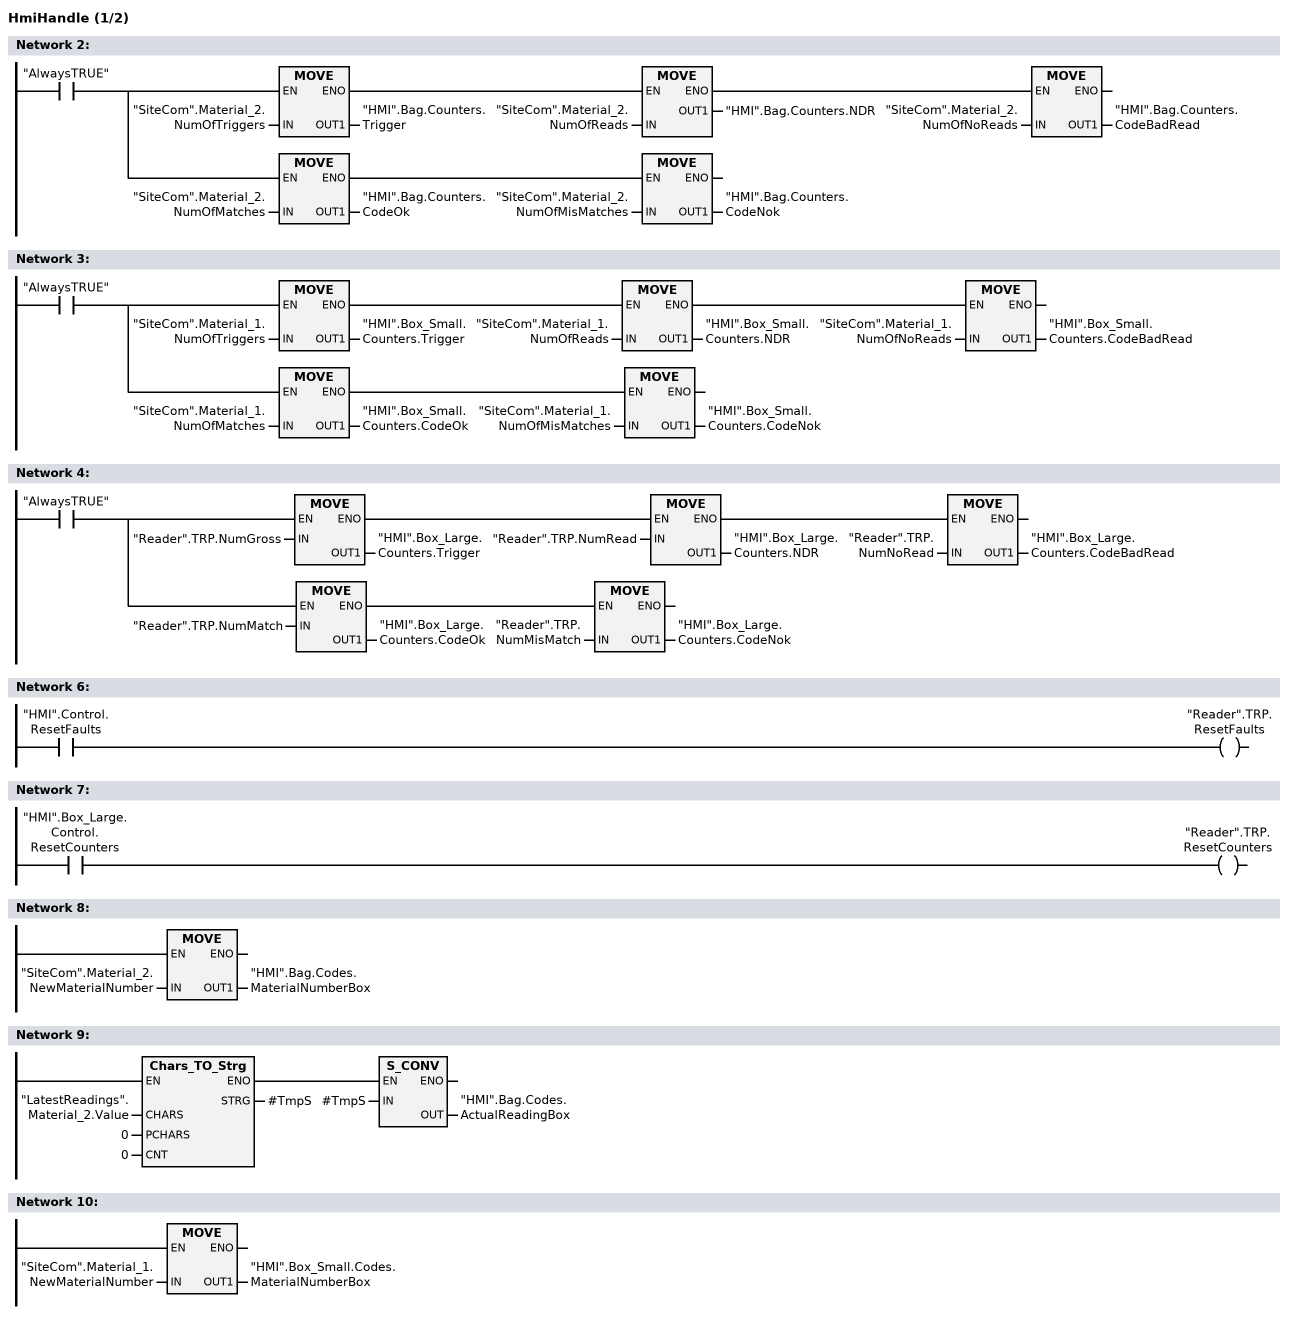
   RUNG wire#powerrail
      Contact( "AlwaysTRUE" )
      wire#w1
      Move(in := "SiteCom".Material_2.NumOfTriggers, out1 => "HMI".Bag.Counters.Trigger)
      Move(in := "SiteCom".Material_2.NumOfReads, out1 => "HMI".Bag.Counters.NDR)
      Move(in := "SiteCom".Material_2.NumOfNoReads, out1 => "HMI".Bag.Counters.CodeBadRead)
   END_RUNG
   RUNG wire#w1
      Move(in := "SiteCom".Material_2.NumOfMatches, out1 => "HMI".Bag.Counters.CodeOk)
      Move(in := "SiteCom".Material_2.NumOfMisMatches, out1 => "HMI".Bag.Counters.CodeNok)
   END_RUNG
   // the same network as SCL:
   IF "AlwaysTRUE" THEN
       "HMI".Bag.Counters.Trigger := "SiteCom".Material_2.NumOfTriggers;
       "HMI".Bag.Counters.NDR := "SiteCom".Material_2.NumOfReads;
       "HMI".Bag.Counters.CodeBadRead := "SiteCom".Material_2.NumOfNoReads;
       "HMI".Bag.Counters.CodeOk := "SiteCom".Material_2.NumOfMatches;
       "HMI".Bag.Counters.CodeNok := "SiteCom".Material_2.NumOfMisMatches;
   END_IF;
END_REGION

REGION Network 3
   RUNG wire#powerrail
      Contact( "AlwaysTRUE" )
      wire#w1
      Move(in := "SiteCom".Material_1.NumOfTriggers, out1 => "HMI".Box_Small.Counters.Trigger)
      Move(in := "SiteCom".Material_1.NumOfReads, out1 => "HMI".Box_Small.Counters.NDR)
      Move(in := "SiteCom".Material_1.NumOfNoReads, out1 => "HMI".Box_Small.Counters.CodeBadRead)
   END_RUNG
   RUNG wire#w1
      Move(in := "SiteCom".Material_1.NumOfMatches, out1 => "HMI".Box_Small.Counters.CodeOk)
      Move(in := "SiteCom".Material_1.NumOfMisMatches, out1 => "HMI".Box_Small.Counters.CodeNok)
   END_RUNG
   // the same network as SCL:
   IF "AlwaysTRUE" THEN
       "HMI".Box_Small.Counters.Trigger := "SiteCom".Material_1.NumOfTriggers;
       "HMI".Box_Small.Counters.NDR := "SiteCom".Material_1.NumOfReads;
       "HMI".Box_Small.Counters.CodeBadRead := "SiteCom".Material_1.NumOfNoReads;
       "HMI".Box_Small.Counters.CodeOk := "SiteCom".Material_1.NumOfMatches;
       "HMI".Box_Small.Counters.CodeNok := "SiteCom".Material_1.NumOfMisMatches;
   END_IF;
END_REGION

REGION Network 4
   RUNG wire#powerrail
      Contact( "AlwaysTRUE" )
      wire#w1
      Move(in := "Reader".TRP.NumGross, out1 => "HMI".Box_Large.Counters.Trigger)
      Move(in := "Reader".TRP.NumRead, out1 => "HMI".Box_Large.Counters.NDR)
      Move(in := "Reader".TRP.NumNoRead, out1 => "HMI".Box_Large.Counters.CodeBadRead)
   END_RUNG
   RUNG wire#w1
      Move(in := "Reader".TRP.NumMatch, out1 => "HMI".Box_Large.Counters.CodeOk)
      Move(in := "Reader".TRP.NumMisMatch, out1 => "HMI".Box_Large.Counters.CodeNok)
   END_RUNG
   // the same network as SCL:
   IF "AlwaysTRUE" THEN
       "HMI".Box_Large.Counters.Trigger := "Reader".TRP.NumGross;
       "HMI".Box_Large.Counters.NDR := "Reader".TRP.NumRead;
       "HMI".Box_Large.Counters.CodeBadRead := "Reader".TRP.NumNoRead;
       "HMI".Box_Large.Counters.CodeOk := "Reader".TRP.NumMatch;
       "HMI".Box_Large.Counters.CodeNok := "Reader".TRP.NumMisMatch;
   END_IF;
END_REGION

REGION Network 6
   RUNG wire#powerrail
      Contact( "HMI".Control.ResetFaults )
      Coil( "Reader".TRP.ResetFaults )
   END_RUNG
   // the same network as SCL:
   "Reader".TRP.ResetFaults := "HMI".Control.ResetFaults;
END_REGION

REGION Network 7
   RUNG wire#powerrail
      Contact( "HMI".Box_Large.Control.ResetCounters )
      Coil( "Reader".TRP.ResetCounters )
   END_RUNG
   // the same network as SCL:
   "Reader".TRP.ResetCounters := "HMI".Box_Large.Control.ResetCounters;
END_REGION

REGION Network 8
   RUNG wire#powerrail
      Move(in := "SiteCom".Material_2.NewMaterialNumber, out1 => "HMI".Bag.Codes.MaterialNumberBox)
   END_RUNG
   // the same network as SCL:
   "HMI".Bag.Codes.MaterialNumberBox := "SiteCom".Material_2.NewMaterialNumber;
END_REGION

REGION Network 9
   // no SCL statement known for Chars_TO_Strg: written as a call
   // ENO of a box is taken as its EN; it also drops when the box reports an error
   Chars_TO_Strg(Chars := "LatestReadings".Material_2.Value, pChars := 0, Cnt := 0, Strg => #TmpS);
   "HMI".Bag.Codes.ActualReadingBox := S_CONV(IN := #TmpS);
END_REGION

REGION Network 10
   RUNG wire#powerrail
      Move(in := "SiteCom".Material_1.NewMaterialNumber, out1 => "HMI".Box_Small.Codes.MaterialNumberBox)
   END_RUNG
   // the same network as SCL:
   "HMI".Box_Small.Codes.MaterialNumberBox := "SiteCom".Material_1.NewMaterialNumber;
END_REGION

REGION Network 11
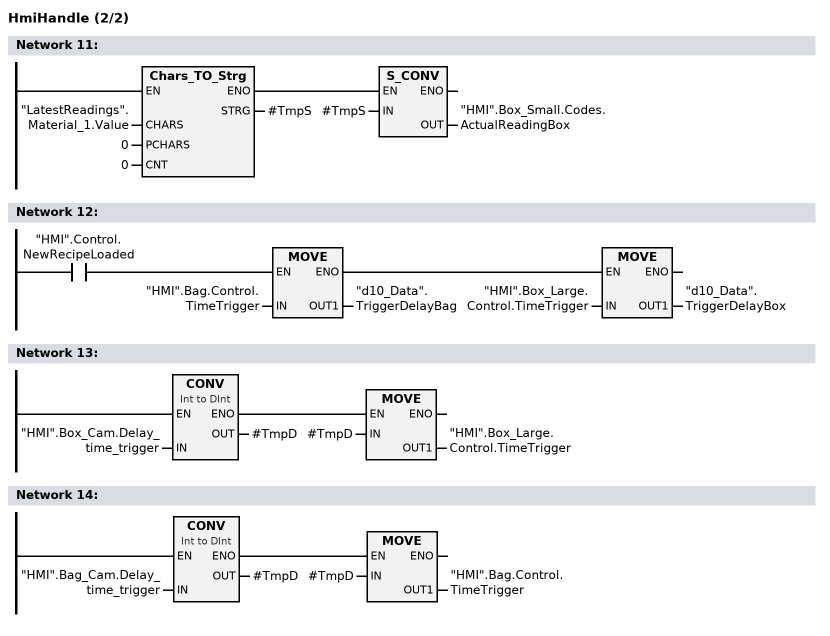
   // no SCL statement known for Chars_TO_Strg: written as a call
   // ENO of a box is taken as its EN; it also drops when the box reports an error
   Chars_TO_Strg(Chars := "LatestReadings".Material_1.Value, pChars := 0, Cnt := 0, Strg => #TmpS);
   "HMI".Box_Small.Codes.ActualReadingBox := S_CONV(IN := #TmpS);
END_REGION

REGION Network 12
   RUNG wire#powerrail
      Contact( "HMI".Control.NewRecipeLoaded )
      Move(in := "HMI".Bag.Control.TimeTrigger, out1 => "d10_Data".TriggerDelayBag)
      Move(in := "HMI".Box_Large.Control.TimeTrigger, out1 => "d10_Data".TriggerDelayBox)
   END_RUNG
   // the same network as SCL:
   IF "HMI".Control.NewRecipeLoaded THEN
       "d10_Data".TriggerDelayBag := "HMI".Bag.Control.TimeTrigger;
       "d10_Data".TriggerDelayBox := "HMI".Box_Large.Control.TimeTrigger;
   END_IF;
END_REGION

REGION Network 13
   RUNG wire#powerrail
      { S7_Templates := "[SrcType := Int, DestType := DInt]" } Convert(in := "HMI".Box_Cam.Delay_time_trigger, out => #TmpD)
      Move(in := #TmpD, out1 => "HMI".Box_Large.Control.TimeTrigger)
   END_RUNG
   // the same network as SCL:
   #TmpD := INT_TO_DINT("HMI".Box_Cam.Delay_time_trigger);
   "HMI".Box_Large.Control.TimeTrigger := #TmpD;
END_REGION

REGION Network 14
   RUNG wire#powerrail
      { S7_Templates := "[SrcType := Int, DestType := DInt]" } Convert(in := "HMI".Bag_Cam.Delay_time_trigger, out => #TmpD)
      Move(in := #TmpD, out1 => "HMI".Bag.Control.TimeTrigger)
   END_RUNG
   // the same network as SCL:
   #TmpD := INT_TO_DINT("HMI".Bag_Cam.Delay_time_trigger);
   "HMI".Bag.Control.TimeTrigger := #TmpD;
END_REGION
END_FUNCTION

FUNCTION "10_DataValidation" : Void   // FC10, LAD
{ S7_Optimized_Access := 'TRUE' }
VERSION : 0.1
BEGIN

REGION Network 1
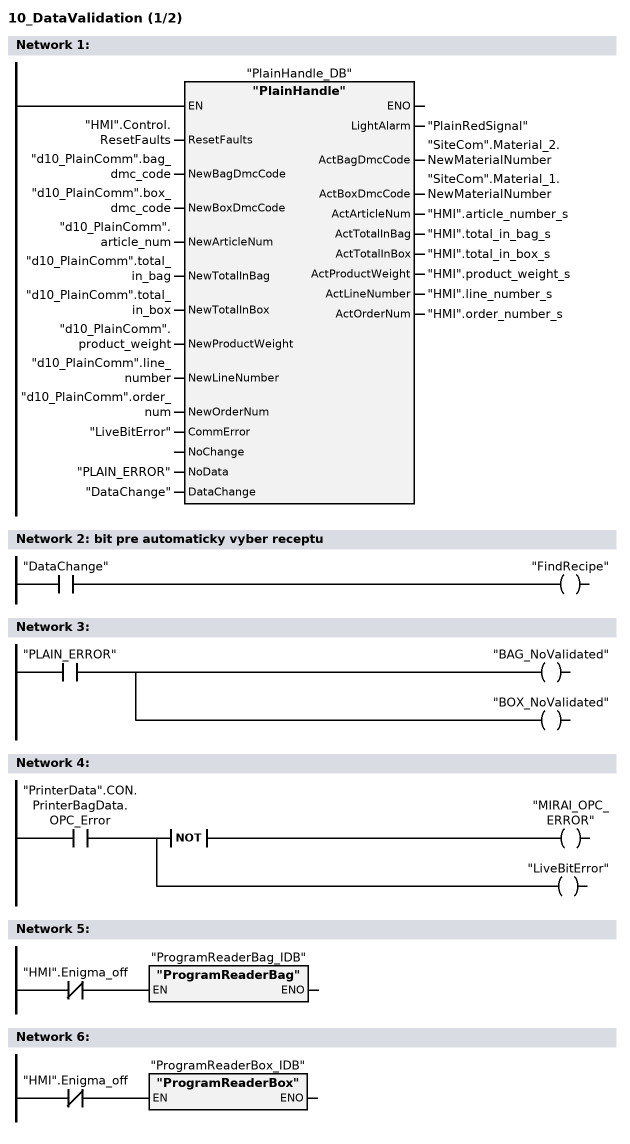
   RUNG wire#powerrail
      "PlainHandle_DB"(ResetFaults := "HMI".Control.ResetFaults, NewBagDmcCode := "d10_PlainComm".bag_dmc_code, NewBoxDmcCode := "d10_PlainComm".box_dmc_code, NewArticleNum := "d10_PlainComm".article_num, NewTotalInBag := "d10_PlainComm".total_in_bag, NewTotalInBox := "d10_PlainComm".total_in_box, NewProductWeight := "d10_PlainComm".product_weight, NewLineNumber := "d10_PlainComm".line_number, NewOrderNum := "d10_PlainComm".order_num, CommError := "LiveBitError", NoChange :=, NoData := "PLAIN_ERROR", DataChange := "DataChange", LightAlarm => "PlainRedSignal", ActBagDmcCode => "SiteCom".Material_2.NewMaterialNumber, ActBoxDmcCode => "SiteCom".Material_1.NewMaterialNumber, ActArticleNum => "HMI".article_number_s, ActTotalInBag => "HMI".total_in_bag_s, ActTotalInBox => "HMI".total_in_box_s, ActProductWeight => "HMI".product_weight_s, ActLineNumber => "HMI".line_number_s, ActOrderNum => "HMI".order_number_s)
   END_RUNG
   // the same network as SCL:
   "PlainHandle_DB"(ResetFaults := "HMI".Control.ResetFaults,   // "PlainHandle"
                    NewBagDmcCode := "d10_PlainComm".bag_dmc_code,
                    NewBoxDmcCode := "d10_PlainComm".box_dmc_code,
                    NewArticleNum := "d10_PlainComm".article_num,
                    NewTotalInBag := "d10_PlainComm".total_in_bag,
                    NewTotalInBox := "d10_PlainComm".total_in_box,
                    NewProductWeight := "d10_PlainComm".product_weight,
                    NewLineNumber := "d10_PlainComm".line_number,
                    NewOrderNum := "d10_PlainComm".order_num,
                    CommError := "LiveBitError",
                    NoData := "PLAIN_ERROR",
                    DataChange := "DataChange",
                    LightAlarm => "PlainRedSignal",
                    ActBagDmcCode => "SiteCom".Material_2.NewMaterialNumber,
                    ActBoxDmcCode => "SiteCom".Material_1.NewMaterialNumber,
                    ActArticleNum => "HMI".article_number_s,
                    ActTotalInBag => "HMI".total_in_bag_s,
                    ActTotalInBox => "HMI".total_in_box_s,
                    ActProductWeight => "HMI".product_weight_s,
                    ActLineNumber => "HMI".line_number_s,
                    ActOrderNum => "HMI".order_number_s);
END_REGION

REGION Network 2: bit pre automaticky vyber receptu
   RUNG wire#powerrail
      Contact( "DataChange" )
      Coil( "FindRecipe" )
   END_RUNG
   // the same network as SCL:
   "FindRecipe" := "DataChange";
END_REGION

REGION Network 3
   RUNG wire#powerrail
      Contact( "PLAIN_ERROR" )
      wire#w1
      Coil( "BAG_NoValidated" )
   END_RUNG
   RUNG wire#w1
      Coil( "BOX_NoValidated" )
   END_RUNG
   // the same network as SCL:
   "BAG_NoValidated" := "PLAIN_ERROR";
   "BOX_NoValidated" := "PLAIN_ERROR";
END_REGION

REGION Network 4
   RUNG wire#powerrail
      Contact( "PrinterData".CON.PrinterBagData.OPC_Error )
      wire#w1
      Not()
      Coil( "MIRAI_OPC_ERROR" )
   END_RUNG
   RUNG wire#w1
      Coil( "LiveBitError" )
   END_RUNG
   // the same network as SCL:
   "MIRAI_OPC_ERROR" := NOT "PrinterData".CON.PrinterBagData.OPC_Error;
   "LiveBitError" := "PrinterData".CON.PrinterBagData.OPC_Error;
END_REGION

REGION Network 5
   RUNG wire#powerrail
      I_Contact( "HMI".Enigma_off )
      "ProgramReaderBag_IDB"()
   END_RUNG
   // the same network as SCL:
   IF NOT "HMI".Enigma_off THEN
       "ProgramReaderBag_IDB"();   // "ProgramReaderBag"
   END_IF;
END_REGION

REGION Network 6
   RUNG wire#powerrail
      I_Contact( "HMI".Enigma_off )
      "ProgramReaderBox_IDB"()
   END_RUNG
   // the same network as SCL:
   IF NOT "HMI".Enigma_off THEN
       "ProgramReaderBox_IDB"();   // "ProgramReaderBox"
   END_IF;
END_REGION

REGION Network 7
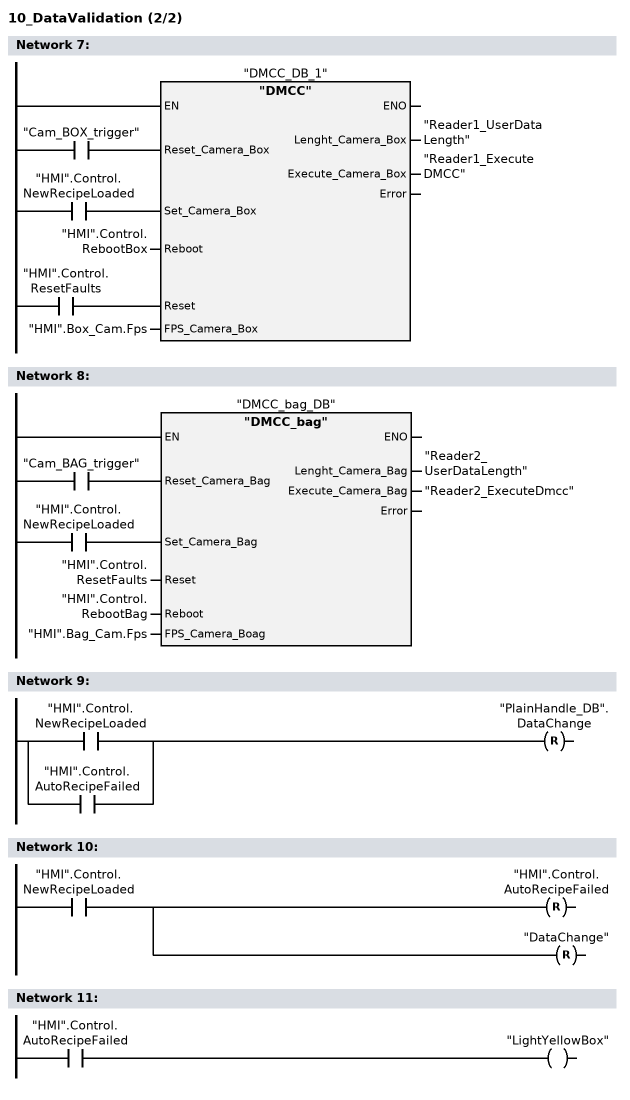
   RUNG wire#powerrail
      "DMCC_DB_1"(Reset_Camera_Box := wire#w1, Set_Camera_Box := wire#w2, Reset := wire#w3, Reboot := "HMI".Control.RebootBox, FPS_Camera_Box := "HMI".Box_Cam.Fps, Lenght_Camera_Box => "Reader1_UserData Length", Execute_Camera_Box => "Reader1_Execute DMCC", Error =>)
   END_RUNG
   RUNG wire#powerrail
      Contact( "Cam_BOX_trigger" )
   END_RUNG wire#w1
   RUNG wire#powerrail
      Contact( "HMI".Control.NewRecipeLoaded )
   END_RUNG wire#w2
   RUNG wire#powerrail
      Contact( "HMI".Control.ResetFaults )
   END_RUNG wire#w3
   // the same network as SCL:
   "DMCC_DB_1"(Reset_Camera_Box := "Cam_BOX_trigger",   // "DMCC"
               Set_Camera_Box := "HMI".Control.NewRecipeLoaded,
               Reboot := "HMI".Control.RebootBox,
               Reset := "HMI".Control.ResetFaults,
               FPS_Camera_Box := "HMI".Box_Cam.Fps,
               Lenght_Camera_Box => "Reader1_UserData Length",
               Execute_Camera_Box => "Reader1_Execute DMCC");
END_REGION

REGION Network 8
   RUNG wire#powerrail
      "DMCC_bag_DB"(Reset_Camera_Bag := wire#w1, Set_Camera_Bag := wire#w2, Reset := "HMI".Control.ResetFaults, Reboot := "HMI".Control.RebootBag, FPS_Camera_Boag := "HMI".Bag_Cam.Fps, Lenght_Camera_Bag => "Reader2_UserDataLength", Execute_Camera_Bag => "Reader2_ExecuteDmcc", Error =>)
   END_RUNG
   RUNG wire#powerrail
      Contact( "Cam_BAG_trigger" )
   END_RUNG wire#w1
   RUNG wire#powerrail
      Contact( "HMI".Control.NewRecipeLoaded )
   END_RUNG wire#w2
   // the same network as SCL:
   "DMCC_bag_DB"(Reset_Camera_Bag := "Cam_BAG_trigger",   // "DMCC_bag"
                 Set_Camera_Bag := "HMI".Control.NewRecipeLoaded,
                 Reset := "HMI".Control.ResetFaults,
                 Reboot := "HMI".Control.RebootBag,
                 FPS_Camera_Boag := "HMI".Bag_Cam.Fps,
                 Lenght_Camera_Bag => "Reader2_UserDataLength",
                 Execute_Camera_Bag => "Reader2_ExecuteDmcc");
END_REGION

REGION Network 9
   RUNG wire#powerrail
      Contact( "HMI".Control.NewRecipeLoaded )
      wire#w1
      R_Coil( "PlainHandle_DB".DataChange )
   END_RUNG
   RUNG wire#powerrail
      Contact( "HMI".Control.AutoRecipeFailed )
   END_RUNG wire#w1
   // the same network as SCL:
   IF "HMI".Control.NewRecipeLoaded OR "HMI".Control.AutoRecipeFailed THEN
       "PlainHandle_DB".DataChange := FALSE;
   END_IF;
END_REGION

REGION Network 10
   RUNG wire#powerrail
      Contact( "HMI".Control.NewRecipeLoaded )
      wire#w1
      R_Coil( "HMI".Control.AutoRecipeFailed )
   END_RUNG
   RUNG wire#w1
      R_Coil( "DataChange" )
   END_RUNG
   // the same network as SCL:
   IF "HMI".Control.NewRecipeLoaded THEN
       "HMI".Control.AutoRecipeFailed := FALSE;
       "DataChange" := FALSE;
   END_IF;
END_REGION

REGION Network 11
   RUNG wire#powerrail
      Contact( "HMI".Control.AutoRecipeFailed )
      Coil( "LightYellowBox" )
   END_RUNG
   // the same network as SCL:
   "LightYellowBox" := "HMI".Control.AutoRecipeFailed;
END_REGION
END_FUNCTION

FUNCTION "20_Mirai" : Void   // FC20, LAD
{ S7_Optimized_Access := 'TRUE' }
VERSION : 0.1
BEGIN

REGION Network 1
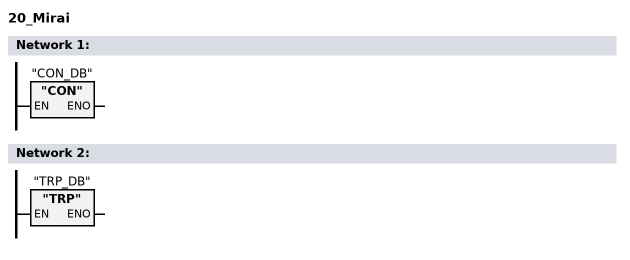
   RUNG wire#powerrail
      "CON_DB"()
   END_RUNG
   // the same network as SCL:
   "CON_DB"();   // "CON"
END_REGION

REGION Network 2
   RUNG wire#powerrail
      "TRP_DB"()
   END_RUNG
   // the same network as SCL:
   "TRP_DB"();   // "TRP"
END_REGION
END_FUNCTION

FUNCTION "FC_CleanQB_Bag" : Void   // FC100, LAD
{ S7_Optimized_Access := 'TRUE' }
VERSION : 0.1
BEGIN

REGION Network 1
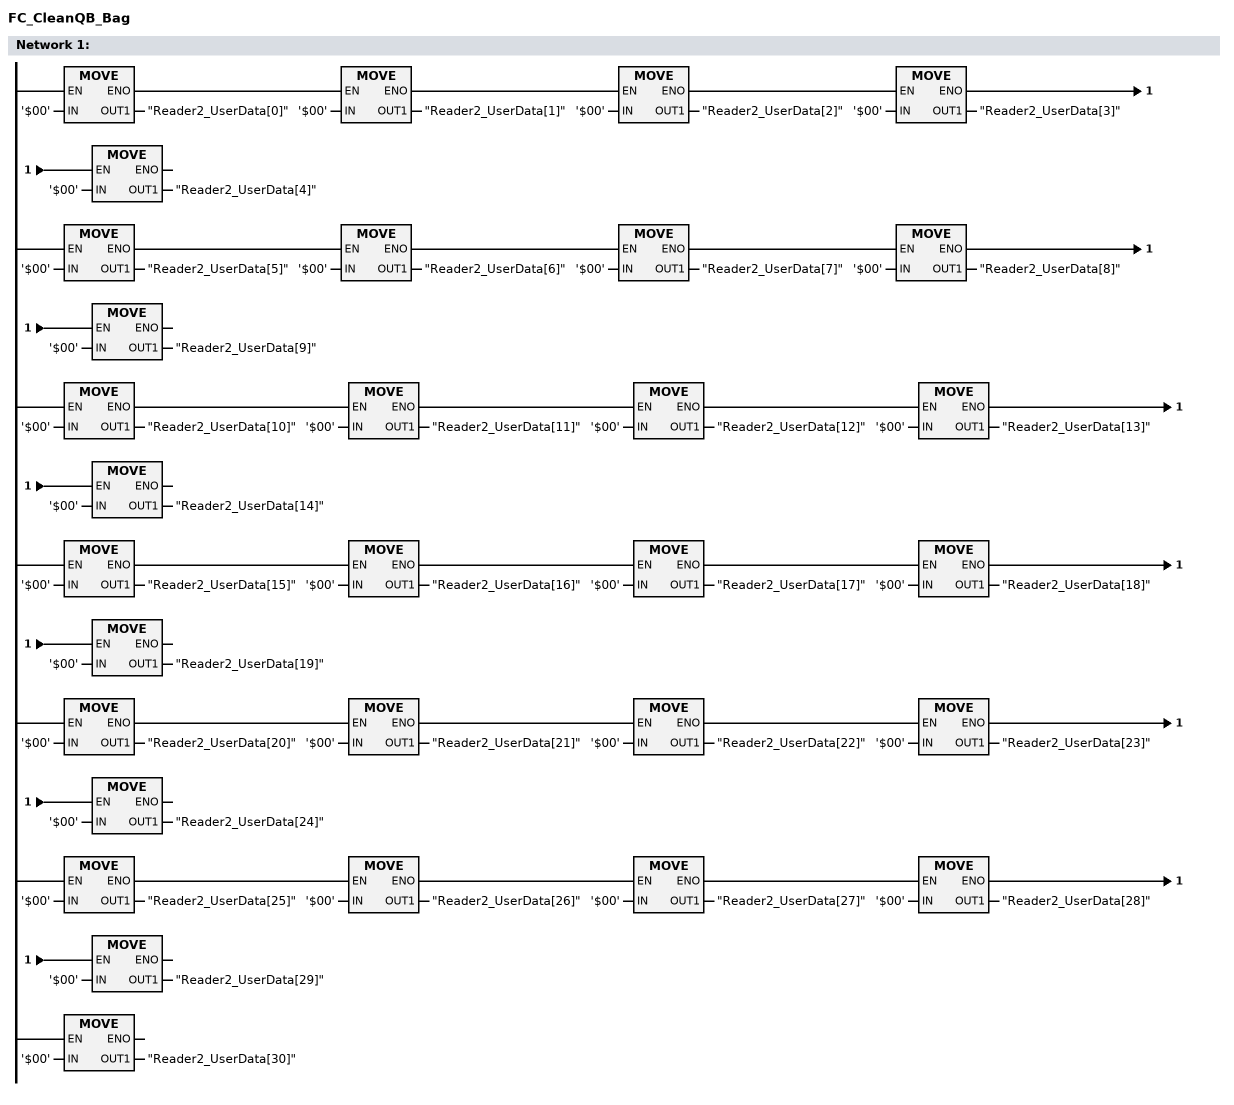
   RUNG wire#powerrail
      Move(in := '$00', out1 => "Reader2_UserData[0]")
      Move(in := '$00', out1 => "Reader2_UserData[1]")
      Move(in := '$00', out1 => "Reader2_UserData[2]")
      Move(in := '$00', out1 => "Reader2_UserData[3]")
      Move(in := '$00', out1 => "Reader2_UserData[4]")
   END_RUNG
   RUNG wire#powerrail
      Move(in := '$00', out1 => "Reader2_UserData[5]")
      Move(in := '$00', out1 => "Reader2_UserData[6]")
      Move(in := '$00', out1 => "Reader2_UserData[7]")
      Move(in := '$00', out1 => "Reader2_UserData[8]")
      Move(in := '$00', out1 => "Reader2_UserData[9]")
   END_RUNG
   RUNG wire#powerrail
      Move(in := '$00', out1 => "Reader2_UserData[10]")
      Move(in := '$00', out1 => "Reader2_UserData[11]")
      Move(in := '$00', out1 => "Reader2_UserData[12]")
      Move(in := '$00', out1 => "Reader2_UserData[13]")
      Move(in := '$00', out1 => "Reader2_UserData[14]")
   END_RUNG
   RUNG wire#powerrail
      Move(in := '$00', out1 => "Reader2_UserData[15]")
      Move(in := '$00', out1 => "Reader2_UserData[16]")
      Move(in := '$00', out1 => "Reader2_UserData[17]")
      Move(in := '$00', out1 => "Reader2_UserData[18]")
      Move(in := '$00', out1 => "Reader2_UserData[19]")
   END_RUNG
   RUNG wire#powerrail
      Move(in := '$00', out1 => "Reader2_UserData[20]")
      Move(in := '$00', out1 => "Reader2_UserData[21]")
      Move(in := '$00', out1 => "Reader2_UserData[22]")
      Move(in := '$00', out1 => "Reader2_UserData[23]")
      Move(in := '$00', out1 => "Reader2_UserData[24]")
   END_RUNG
   RUNG wire#powerrail
      Move(in := '$00', out1 => "Reader2_UserData[25]")
      Move(in := '$00', out1 => "Reader2_UserData[26]")
      Move(in := '$00', out1 => "Reader2_UserData[27]")
      Move(in := '$00', out1 => "Reader2_UserData[28]")
      Move(in := '$00', out1 => "Reader2_UserData[29]")
   END_RUNG
   RUNG wire#powerrail
      Move(in := '$00', out1 => "Reader2_UserData[30]")
   END_RUNG
   // the same network as SCL:
   "Reader2_UserData[0]" := '$00';
   "Reader2_UserData[1]" := '$00';
   "Reader2_UserData[2]" := '$00';
   "Reader2_UserData[3]" := '$00';
   "Reader2_UserData[4]" := '$00';
   "Reader2_UserData[5]" := '$00';
   "Reader2_UserData[6]" := '$00';
   "Reader2_UserData[7]" := '$00';
   "Reader2_UserData[8]" := '$00';
   "Reader2_UserData[9]" := '$00';
   "Reader2_UserData[10]" := '$00';
   "Reader2_UserData[11]" := '$00';
   "Reader2_UserData[12]" := '$00';
   "Reader2_UserData[13]" := '$00';
   "Reader2_UserData[14]" := '$00';
   "Reader2_UserData[15]" := '$00';
   "Reader2_UserData[16]" := '$00';
   "Reader2_UserData[17]" := '$00';
   "Reader2_UserData[18]" := '$00';
   "Reader2_UserData[19]" := '$00';
   "Reader2_UserData[20]" := '$00';
   "Reader2_UserData[21]" := '$00';
   "Reader2_UserData[22]" := '$00';
   "Reader2_UserData[23]" := '$00';
   "Reader2_UserData[24]" := '$00';
   "Reader2_UserData[25]" := '$00';
   "Reader2_UserData[26]" := '$00';
   "Reader2_UserData[27]" := '$00';
   "Reader2_UserData[28]" := '$00';
   "Reader2_UserData[29]" := '$00';
   "Reader2_UserData[30]" := '$00';
END_REGION
END_FUNCTION

FUNCTION "FC_CleanQB_Box" : Void   // FC101, LAD
{ S7_Optimized_Access := 'TRUE' }
VERSION : 0.1
BEGIN

REGION Network 1
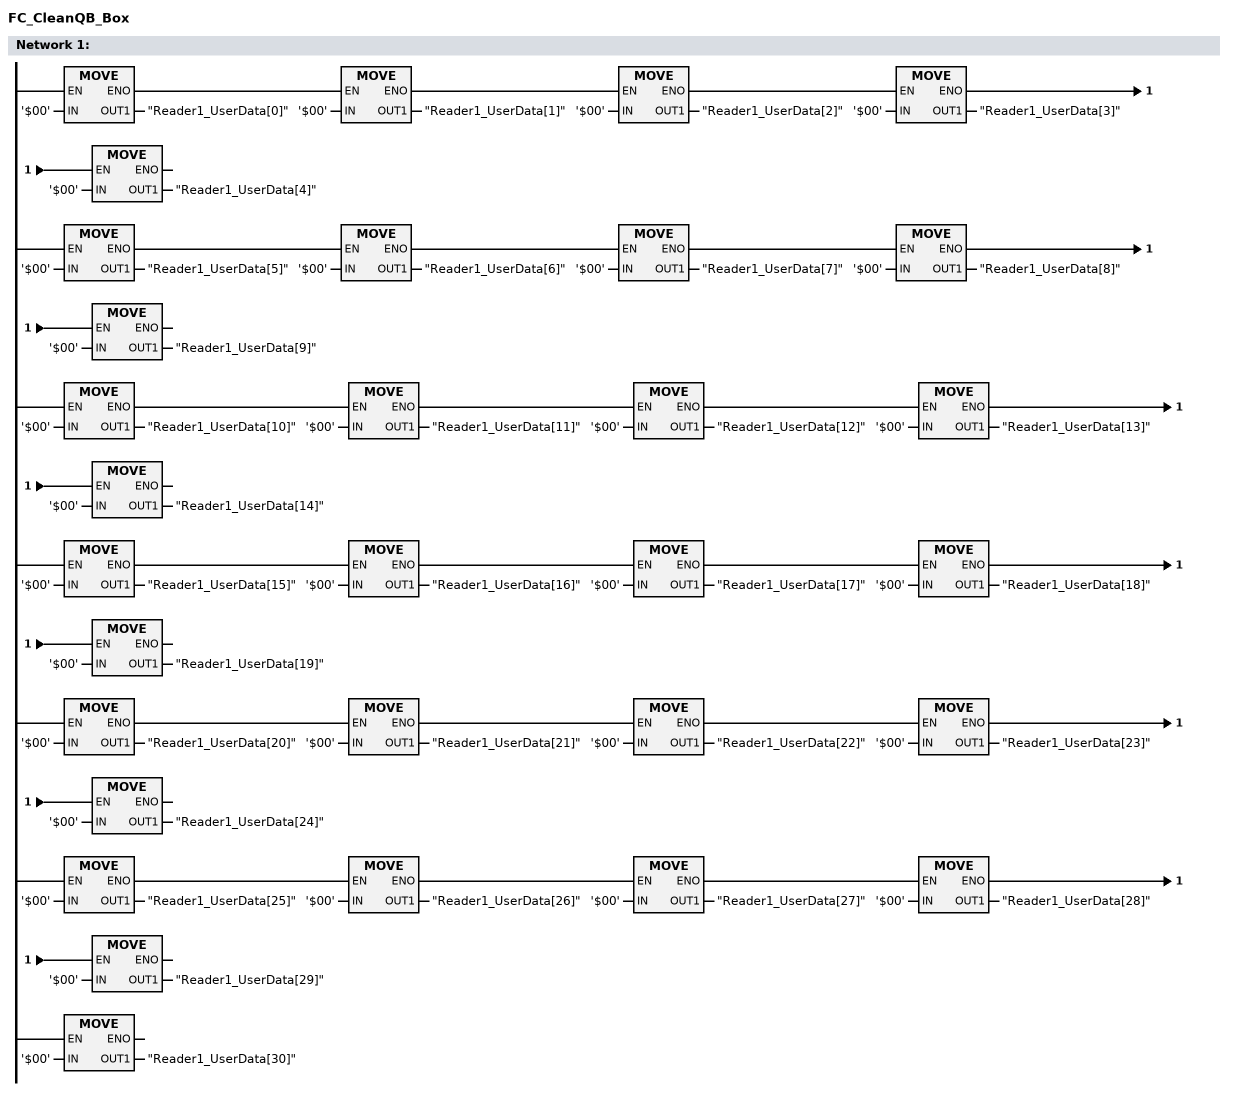
   RUNG wire#powerrail
      Move(in := '$00', out1 => "Reader1_UserData[0]")
      Move(in := '$00', out1 => "Reader1_UserData[1]")
      Move(in := '$00', out1 => "Reader1_UserData[2]")
      Move(in := '$00', out1 => "Reader1_UserData[3]")
      Move(in := '$00', out1 => "Reader1_UserData[4]")
   END_RUNG
   RUNG wire#powerrail
      Move(in := '$00', out1 => "Reader1_UserData[5]")
      Move(in := '$00', out1 => "Reader1_UserData[6]")
      Move(in := '$00', out1 => "Reader1_UserData[7]")
      Move(in := '$00', out1 => "Reader1_UserData[8]")
      Move(in := '$00', out1 => "Reader1_UserData[9]")
   END_RUNG
   RUNG wire#powerrail
      Move(in := '$00', out1 => "Reader1_UserData[10]")
      Move(in := '$00', out1 => "Reader1_UserData[11]")
      Move(in := '$00', out1 => "Reader1_UserData[12]")
      Move(in := '$00', out1 => "Reader1_UserData[13]")
      Move(in := '$00', out1 => "Reader1_UserData[14]")
   END_RUNG
   RUNG wire#powerrail
      Move(in := '$00', out1 => "Reader1_UserData[15]")
      Move(in := '$00', out1 => "Reader1_UserData[16]")
      Move(in := '$00', out1 => "Reader1_UserData[17]")
      Move(in := '$00', out1 => "Reader1_UserData[18]")
      Move(in := '$00', out1 => "Reader1_UserData[19]")
   END_RUNG
   RUNG wire#powerrail
      Move(in := '$00', out1 => "Reader1_UserData[20]")
      Move(in := '$00', out1 => "Reader1_UserData[21]")
      Move(in := '$00', out1 => "Reader1_UserData[22]")
      Move(in := '$00', out1 => "Reader1_UserData[23]")
      Move(in := '$00', out1 => "Reader1_UserData[24]")
   END_RUNG
   RUNG wire#powerrail
      Move(in := '$00', out1 => "Reader1_UserData[25]")
      Move(in := '$00', out1 => "Reader1_UserData[26]")
      Move(in := '$00', out1 => "Reader1_UserData[27]")
      Move(in := '$00', out1 => "Reader1_UserData[28]")
      Move(in := '$00', out1 => "Reader1_UserData[29]")
   END_RUNG
   RUNG wire#powerrail
      Move(in := '$00', out1 => "Reader1_UserData[30]")
   END_RUNG
   // the same network as SCL:
   "Reader1_UserData[0]" := '$00';
   "Reader1_UserData[1]" := '$00';
   "Reader1_UserData[2]" := '$00';
   "Reader1_UserData[3]" := '$00';
   "Reader1_UserData[4]" := '$00';
   "Reader1_UserData[5]" := '$00';
   "Reader1_UserData[6]" := '$00';
   "Reader1_UserData[7]" := '$00';
   "Reader1_UserData[8]" := '$00';
   "Reader1_UserData[9]" := '$00';
   "Reader1_UserData[10]" := '$00';
   "Reader1_UserData[11]" := '$00';
   "Reader1_UserData[12]" := '$00';
   "Reader1_UserData[13]" := '$00';
   "Reader1_UserData[14]" := '$00';
   "Reader1_UserData[15]" := '$00';
   "Reader1_UserData[16]" := '$00';
   "Reader1_UserData[17]" := '$00';
   "Reader1_UserData[18]" := '$00';
   "Reader1_UserData[19]" := '$00';
   "Reader1_UserData[20]" := '$00';
   "Reader1_UserData[21]" := '$00';
   "Reader1_UserData[22]" := '$00';
   "Reader1_UserData[23]" := '$00';
   "Reader1_UserData[24]" := '$00';
   "Reader1_UserData[25]" := '$00';
   "Reader1_UserData[26]" := '$00';
   "Reader1_UserData[27]" := '$00';
   "Reader1_UserData[28]" := '$00';
   "Reader1_UserData[29]" := '$00';
   "Reader1_UserData[30]" := '$00';
END_REGION
END_FUNCTION

FUNCTION "LGF_StringToTaddr" : TADDR_Param   // FC10041, SCL
{ S7_Optimized_Access := 'TRUE' }
VERSION : 0.1
   VAR_INPUT
      ipAddressString : String;
   END_VAR
   VAR_OUTPUT
      error : Bool;
      status : Word;
   END_VAR
   VAR_TEMP
      tempCharPosition : Int;
      tempAddressString : String;
      tempOctetString : String[4];
      tempUInt : UInt;
      tempPortNumberIsSpecified : Bool;
      tempIpAdressTaddr : TADDR_Param;
   END_VAR
   VAR CONSTANT
      NO_ERROR : Word := 16#0000;
      WRONG_VALUE_POS1 : Word := 16#8101;
      WRONG_VALUE_POS2 : Word := 16#8102;
      WRONG_VALUE_POS3 : Word := 16#8103;
      WRONG_VALUE_POS4 : Word := 16#8104;
      WRONG_VALUE_PORT : Word := 16#8105;
      MAX_USINT : USInt := 255;
      MAX_UINT : UInt := 65535;
      EMPTY_STRING : String := '';
      MAX_CHAR_FOR_IP_PART : Int := 4;
      MAX_CHAR_FOR_PORT_PART : Int := 5;
      INIT_VAL : USInt := 0;
      NO_POS : Int := 0;
   END_VAR
BEGIN
   //=============================================================================
   // SIEMENS AG
   // (c)Copyright 2017
   //-----------------------------------------------------------------------------
   // Library:       LGF (Library General Functions)
   // Tested with:   CPU1212C DC/DC/DC FW:V4.2
   // Engineering:   TIA Portal V14 Upd 1
   // Restrictions:  -
   // Requirements:  PLC (S7-1200 / S7-1500)
   // Functionality: This function converts a string IP Address
   //                into TADDR Param format.
   //-----------------------------------------------------------------------------
   // Change log table:
   // Version  Date       In charge Changes applied
   // 01.00.00 30.01.2017 Siemens Industry Online Support
   //                     First released version
   //-----------------------------------------------------------------------------
   //Status Codes:
   // 16#0000:  No errors
   // 16#8101:  Wrong value on position 1
   // 16#8102:  Wrong value on position 2
   // 16#8103:  Wrong value on position 3
   // 16#8104:  Wrong value on position 4
   // 16#8105:  Wrong value on port position
   //=============================================================================

   // Initialization
   #error := FALSE;
   #status := #NO_ERROR;
   #tempAddressString := #ipAddressString;
   #LGF_StringToTaddr.REM_IP_ADDR[1] := #INIT_VAL;
   #LGF_StringToTaddr.REM_IP_ADDR[2] := #INIT_VAL;
   #LGF_StringToTaddr.REM_IP_ADDR[3] := #INIT_VAL;
   #LGF_StringToTaddr.REM_IP_ADDR[4] := #INIT_VAL;
   #LGF_StringToTaddr.REM_PORT_NR := #INIT_VAL;

   // Process the 1st octet of the IP Address
   #tempCharPosition := FIND(IN1 := #tempAddressString, IN2 := '.');
   IF #tempCharPosition > #MAX_CHAR_FOR_IP_PART THEN
     #error := TRUE;
     #status := #WRONG_VALUE_POS1;
     RETURN;
   ELSE
     #tempOctetString := LEFT(IN := #tempAddressString, L := #tempCharPosition - 1);
     // Check if string is empty
     IF #tempOctetString = #EMPTY_STRING THEN
       #error := TRUE;
       #status := #WRONG_VALUE_POS1;
       RETURN;
     ELSE
       #tempAddressString := DELETE(IN := #tempAddressString, P := 1, L := #tempCharPosition);
     END_IF;
   END_IF;

   // Convert the 1st octet string to numerical value
   STRG_VAL(IN := #tempOctetString,
            FORMAT := W#16#0000,
            P := 1,
            OUT => #tempUInt);

     IF #tempUInt > #MAX_USINT THEN
       #error := TRUE;
       #status := #WRONG_VALUE_POS1;
       RETURN;
     ELSE
       #tempIpAdressTaddr.REM_IP_ADDR[1] := UINT_TO_BYTE(#tempUInt);
     END_IF;


   // Process the 2nd octetstring of the IP Address
   #tempCharPosition := FIND(IN1 := #tempAddressString, IN2 := '.');
   IF #tempCharPosition > #MAX_CHAR_FOR_IP_PART THEN
     #error := TRUE;
     #status := #WRONG_VALUE_POS2;
     RETURN;
   ELSE
     #tempOctetString := LEFT(IN := #tempAddressString, L := #tempCharPosition - 1);
     IF #tempOctetString = #EMPTY_STRING THEN
       #error := TRUE;
       #status := #WRONG_VALUE_POS2;
       RETURN;
     ELSE
       #tempAddressString := DELETE(IN := #tempAddressString, P := 1, L := #tempCharPosition);
     END_IF;
   END_IF;

   // Convert the 2nd octet string TO numerical value
   STRG_VAL(IN := #tempOctetString,
            FORMAT := W#16#0000,
            P := 1,
            OUT => #tempUInt);

   IF #tempUInt > #MAX_USINT THEN
     #error := TRUE;
     #status := #WRONG_VALUE_POS2;
     RETURN;
   ELSE
     #tempIpAdressTaddr.REM_IP_ADDR[2] := UINT_TO_BYTE(#tempUInt);
   END_IF;

   // Process the 3rd octet of the IP Address
   #tempCharPosition := FIND(IN1 := #tempAddressString, IN2 := '.');
   IF #tempCharPosition > #MAX_CHAR_FOR_IP_PART THEN
     #error := TRUE;
     #status := #WRONG_VALUE_POS3;
     RETURN;
   ELSE
     #tempOctetString := LEFT(IN := #tempAddressString, L := #tempCharPosition - 1);
     // Check if string is empty
     IF #tempOctetString = #EMPTY_STRING THEN
       #error := TRUE;
       #status := #WRONG_VALUE_POS3;
       RETURN;
     ELSE
       #tempAddressString := DELETE(IN := #tempAddressString, P := 1, L := #tempCharPosition);
     END_IF;
   END_IF;